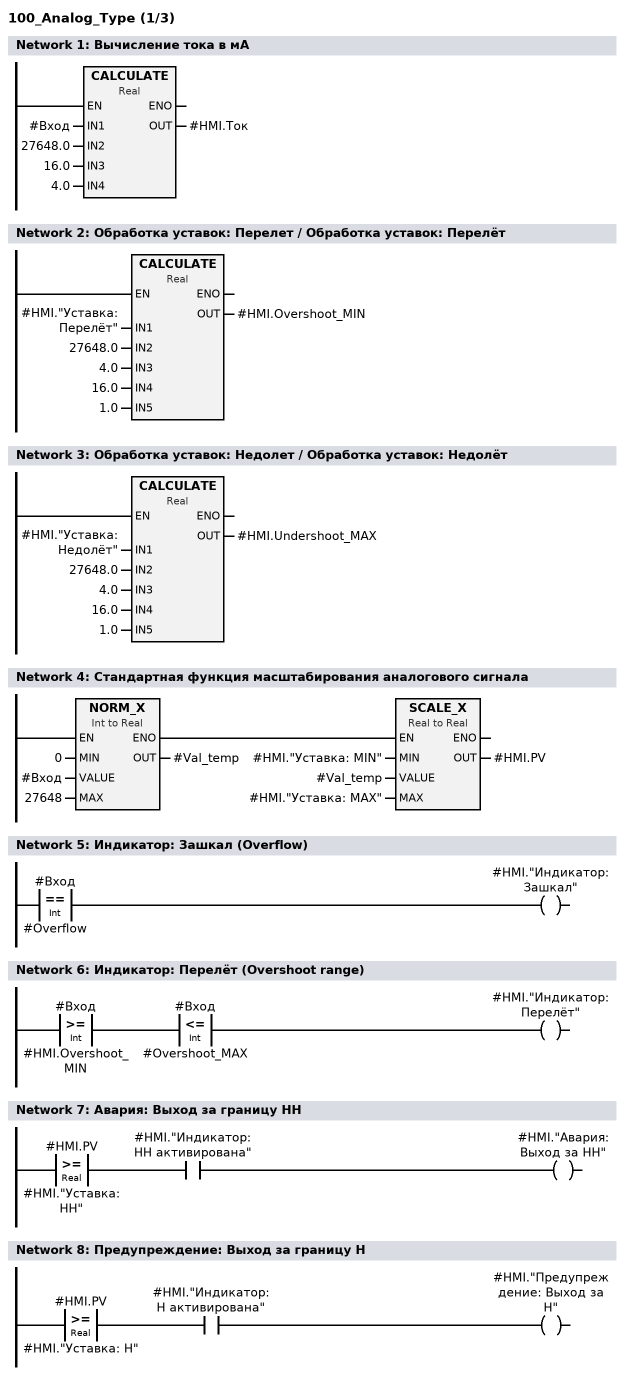
   RUNG wire#powerrail
      { S7_Templates := "SrcType := Real"; S7_Expression := "((IN3 / IN2) * IN1 + IN4)" } Calculate(in1 := #Вход, in2 := 27648.0, in3 := 16.0, in4 := 4.0, out => #HMI.Ток)
   END_RUNG
   // the same network as SCL:
   #HMI.Ток := ((16.0 / 27648.0) * #Вход + 4.0);
END_REGION

REGION Network 2: Обработка уставок: Перелет / Обработка уставок: Перелёт
   RUNG wire#powerrail
      { S7_Templates := "SrcType := Real"; S7_Expression := "((IN1- IN3) * IN2 / IN4) +IN5" } Calculate(in1 := #HMI."Уставка: Перелёт", in2 := 27648.0, in3 := 4.0, in4 := 16.0, in5 := 1.0, out => #HMI.Overshoot_MIN)
   END_RUNG
   // the same network as SCL:
   #HMI.Overshoot_MIN := ((#HMI."Уставка: Перелёт"- 4.0) * 27648.0 / 16.0) +1.0;
END_REGION

REGION Network 3: Обработка уставок: Недолет / Обработка уставок: Недолёт
   RUNG wire#powerrail
      { S7_Templates := "SrcType := Real"; S7_Expression := "((IN1- IN3) * IN2 / IN4) - IN5" } Calculate(in1 := #HMI."Уставка: Недолёт", in2 := 27648.0, in3 := 4.0, in4 := 16.0, in5 := 1.0, out => #HMI.Undershoot_MAX)
   END_RUNG
   // the same network as SCL:
   #HMI.Undershoot_MAX := ((#HMI."Уставка: Недолёт"- 4.0) * 27648.0 / 16.0) - 1.0;
END_REGION

REGION Network 4: Стандартная функция масштабирования аналогового сигнала
   RUNG wire#powerrail
      { S7_Templates := "[SrcType := Int, DestType := Real]" } Normalize(min := 0, value := #Вход, max := 27648, out => #Val_temp)
      { S7_Templates := "[SrcType := Real, DestType := Real]" } Scale(min := #HMI."Уставка: MIN", value := #Val_temp, max := #HMI."Уставка: MAX", out => #HMI.PV)
   END_RUNG
   // the same network as SCL:
   #Val_temp := NORM_X(MIN := 0, VALUE := #Вход, MAX := 27648);
   #HMI.PV := SCALE_X(MIN := #HMI."Уставка: MIN", VALUE := #Val_temp, MAX := #HMI."Уставка: MAX");
END_REGION

REGION Network 5: Индикатор: Зашкал (Overflow)
   RUNG wire#powerrail
      { S7_Templates := "SrcType := Int" } EQ_Contact(in1 := #Вход, in2 := #Overflow)
      Coil( #HMI."Индикатор: Зашкал" )
   END_RUNG
   // the same network as SCL:
   #HMI."Индикатор: Зашкал" := #Вход = #Overflow;
END_REGION

REGION Network 6: Индикатор: Перелёт (Overshoot range)
   RUNG wire#powerrail
      { S7_Templates := "SrcType := Int" } GE_Contact(in1 := #Вход, in2 := #HMI.Overshoot_MIN)
      { S7_Templates := "SrcType := Int" } LE_Contact(in1 := #Вход, in2 := #Overshoot_MAX)
      Coil( #HMI."Индикатор: Перелёт" )
   END_RUNG
   // the same network as SCL:
   #HMI."Индикатор: Перелёт" := (#Вход >= #HMI.Overshoot_MIN) AND (#Вход <= #Overshoot_MAX);
END_REGION

REGION Network 7: Авария: Выход за границу НН
   RUNG wire#powerrail
      { S7_Templates := "SrcType := Real" } GE_Contact(in1 := #HMI.PV, in2 := #HMI."Уставка: HH")
      Contact( #HMI."Индикатор: HH активирована" )
      Coil( #HMI."Авария: Выход за HH" )
   END_RUNG
   // the same network as SCL:
   #HMI."Авария: Выход за HH" := (#HMI.PV >= #HMI."Уставка: HH") AND #HMI."Индикатор: HH активирована";
END_REGION

REGION Network 8: Предупреждение: Выход за границу Н
   RUNG wire#powerrail
      { S7_Templates := "SrcType := Real" } GE_Contact(in1 := #HMI.PV, in2 := #HMI."Уставка: H")
      Contact( #HMI."Индикатор: H активирована" )
      Coil( #HMI."Предупреждение: Выход за H" )
   END_RUNG
   // the same network as SCL:
   #HMI."Предупреждение: Выход за H" := (#HMI.PV >= #HMI."Уставка: H") AND #HMI."Индикатор: H активирована";
END_REGION

REGION Network 9: Предупреждение: Выход за границу L
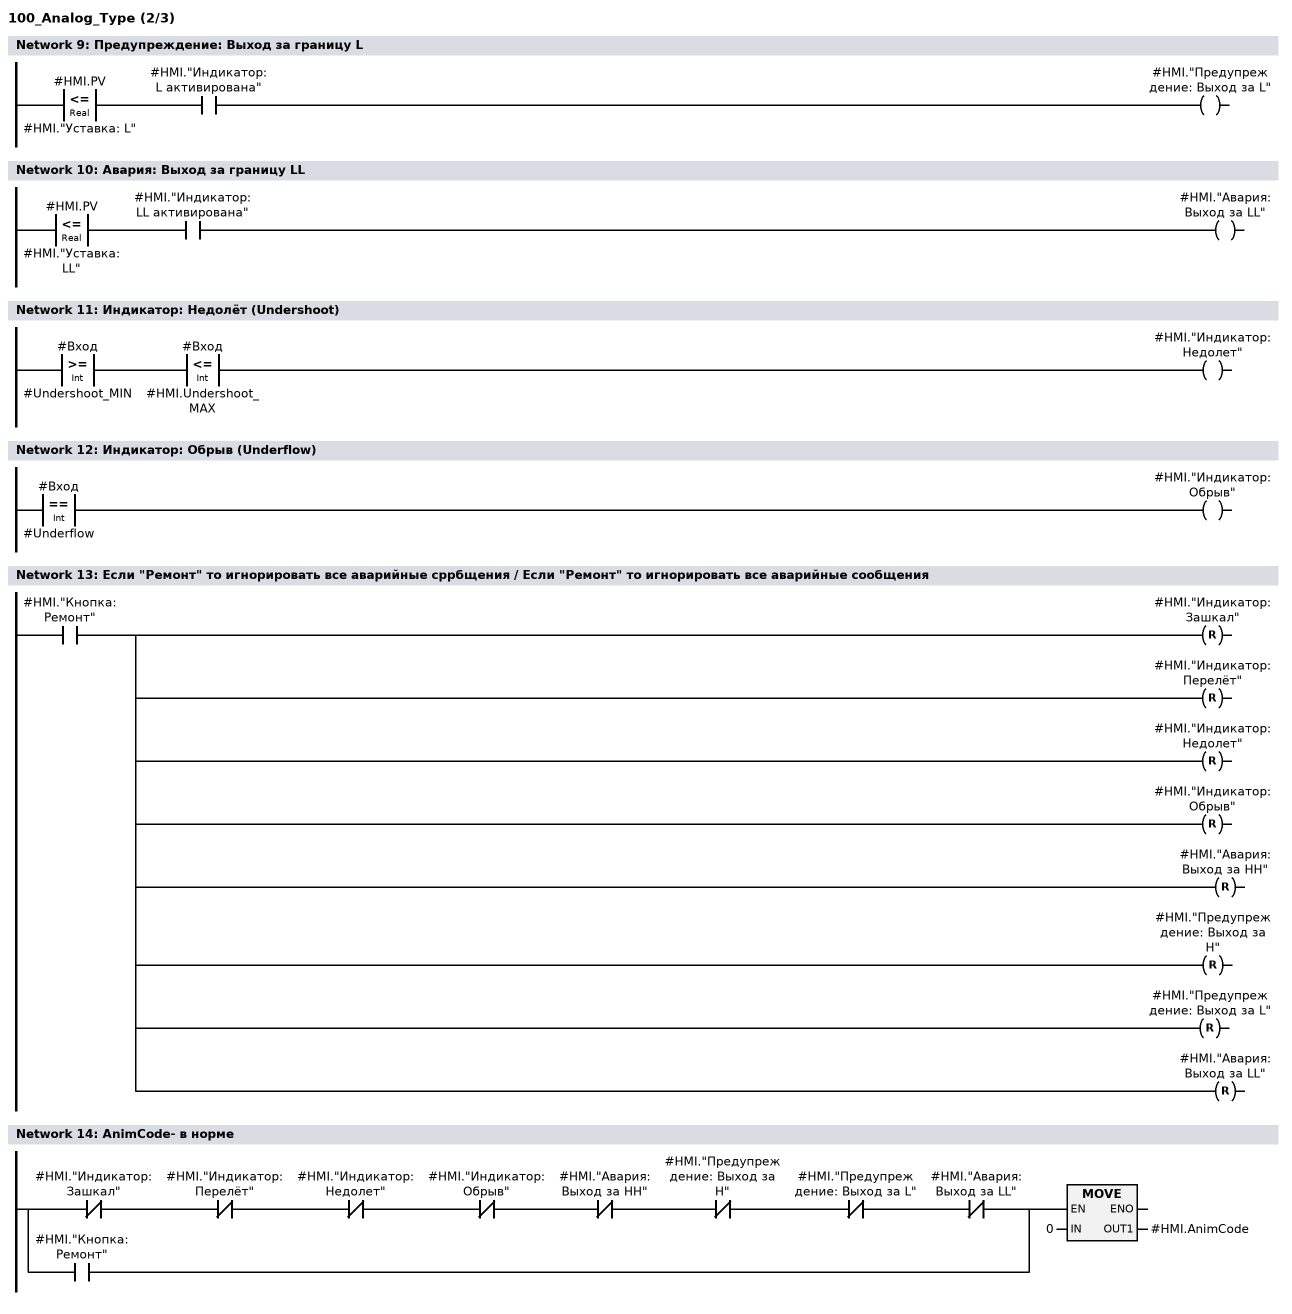
   RUNG wire#powerrail
      { S7_Templates := "SrcType := Real" } LE_Contact(in1 := #HMI.PV, in2 := #HMI."Уставка: L")
      Contact( #HMI."Индикатор: L активирована" )
      Coil( #HMI."Предупреждение: Выход за L" )
   END_RUNG
   // the same network as SCL:
   #HMI."Предупреждение: Выход за L" := (#HMI.PV <= #HMI."Уставка: L") AND #HMI."Индикатор: L активирована";
END_REGION

REGION Network 10: Авария: Выход за границу LL
   RUNG wire#powerrail
      { S7_Templates := "SrcType := Real" } LE_Contact(in1 := #HMI.PV, in2 := #HMI."Уставка: LL")
      Contact( #HMI."Индикатор: LL активирована" )
      Coil( #HMI."Авария: Выход за LL" )
   END_RUNG
   // the same network as SCL:
   #HMI."Авария: Выход за LL" := (#HMI.PV <= #HMI."Уставка: LL") AND #HMI."Индикатор: LL активирована";
END_REGION

REGION Network 11: Индикатор: Недолёт (Undershoot)
   RUNG wire#powerrail
      { S7_Templates := "SrcType := Int" } GE_Contact(in1 := #Вход, in2 := #Undershoot_MIN)
      { S7_Templates := "SrcType := Int" } LE_Contact(in1 := #Вход, in2 := #HMI.Undershoot_MAX)
      Coil( #HMI."Индикатор: Недолет" )
   END_RUNG
   // the same network as SCL:
   #HMI."Индикатор: Недолет" := (#Вход >= #Undershoot_MIN) AND (#Вход <= #HMI.Undershoot_MAX);
END_REGION

REGION Network 12: Индикатор: Обрыв (Underflow)
   RUNG wire#powerrail
      { S7_Templates := "SrcType := Int" } EQ_Contact(in1 := #Вход, in2 := #Underflow)
      Coil( #HMI."Индикатор: Обрыв" )
   END_RUNG
   // the same network as SCL:
   #HMI."Индикатор: Обрыв" := #Вход = #Underflow;
END_REGION

REGION Network 13: Если "Ремонт" то игнорировать все аварийные сррбщения / Если "Ремонт" то игнорировать все аварийные сообщения
   RUNG wire#powerrail
      Contact( #HMI."Кнопка: Ремонт" )
      wire#w1
      R_Coil( #HMI."Индикатор: Зашкал" )
   END_RUNG
   RUNG wire#w1
      R_Coil( #HMI."Индикатор: Перелёт" )
   END_RUNG
   RUNG wire#w1
      R_Coil( #HMI."Индикатор: Недолет" )
   END_RUNG
   RUNG wire#w1
      R_Coil( #HMI."Индикатор: Обрыв" )
   END_RUNG
   RUNG wire#w1
      R_Coil( #HMI."Авария: Выход за HH" )
   END_RUNG
   RUNG wire#w1
      R_Coil( #HMI."Предупреждение: Выход за H" )
   END_RUNG
   RUNG wire#w1
      R_Coil( #HMI."Предупреждение: Выход за L" )
   END_RUNG
   RUNG wire#w1
      R_Coil( #HMI."Авария: Выход за LL" )
   END_RUNG
   // the same network as SCL:
   IF #HMI."Кнопка: Ремонт" THEN
       #HMI."Индикатор: Зашкал" := FALSE;
       #HMI."Индикатор: Перелёт" := FALSE;
       #HMI."Индикатор: Недолет" := FALSE;
       #HMI."Индикатор: Обрыв" := FALSE;
       #HMI."Авария: Выход за HH" := FALSE;
       #HMI."Предупреждение: Выход за H" := FALSE;
       #HMI."Предупреждение: Выход за L" := FALSE;
       #HMI."Авария: Выход за LL" := FALSE;
   END_IF;
END_REGION

REGION Network 14: AnimCode- в норме
   RUNG wire#powerrail
      I_Contact( #HMI."Индикатор: Зашкал" )
      I_Contact( #HMI."Индикатор: Перелёт" )
      I_Contact( #HMI."Индикатор: Недолет" )
      I_Contact( #HMI."Индикатор: Обрыв" )
      I_Contact( #HMI."Авария: Выход за HH" )
      I_Contact( #HMI."Предупреждение: Выход за H" )
      I_Contact( #HMI."Предупреждение: Выход за L" )
      I_Contact( #HMI."Авария: Выход за LL" )
      wire#w1
      Move(in := 0, out1 => #HMI.AnimCode)
   END_RUNG
   RUNG wire#powerrail
      Contact( #HMI."Кнопка: Ремонт" )
   END_RUNG wire#w1
   // the same network as SCL:
   IF (NOT #HMI."Индикатор: Зашкал" AND NOT #HMI."Индикатор: Перелёт" AND NOT #HMI."Индикатор: Недолет" AND NOT #HMI."Индикатор: Обрыв" AND NOT #HMI."Авария: Выход за HH" AND NOT #HMI."Предупреждение: Выход за H" AND NOT #HMI."Предупреждение: Выход за L" AND NOT #HMI."Авария: Выход за LL") OR #HMI."Кнопка: Ремонт" THEN
       #HMI.AnimCode := 0;
   END_IF;
END_REGION

REGION Network 15: AnimCode- предупреждение
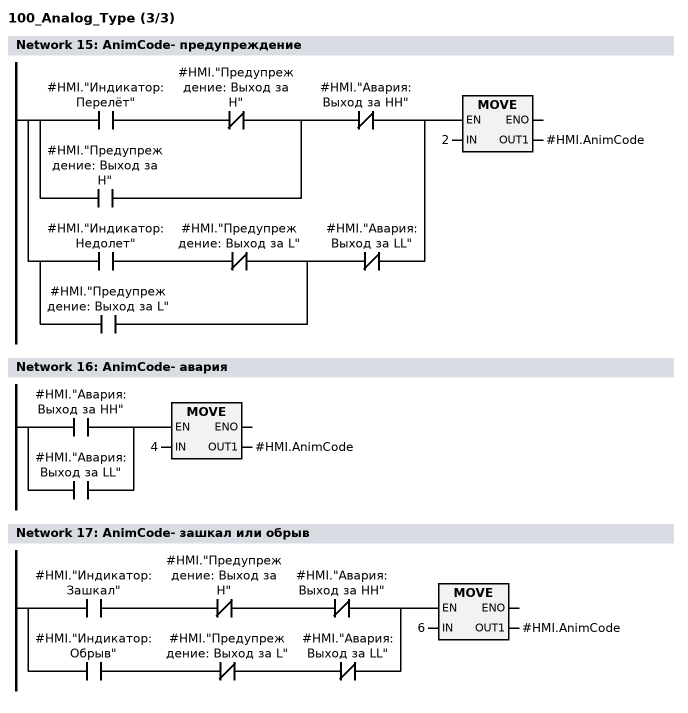
   RUNG wire#powerrail
      Contact( #HMI."Индикатор: Перелёт" )
      I_Contact( #HMI."Предупреждение: Выход за H" )
      wire#w1
      I_Contact( #HMI."Авария: Выход за HH" )
      wire#w2
      Move(in := 2, out1 => #HMI.AnimCode)
   END_RUNG
   RUNG wire#powerrail
      Contact( #HMI."Предупреждение: Выход за H" )
   END_RUNG wire#w1
   RUNG wire#powerrail
      Contact( #HMI."Индикатор: Недолет" )
      I_Contact( #HMI."Предупреждение: Выход за L" )
      wire#w3
      I_Contact( #HMI."Авария: Выход за LL" )
   END_RUNG wire#w2
   RUNG wire#powerrail
      Contact( #HMI."Предупреждение: Выход за L" )
   END_RUNG wire#w3
   // the same network as SCL:
   IF (((#HMI."Индикатор: Перелёт" AND NOT #HMI."Предупреждение: Выход за H") OR #HMI."Предупреждение: Выход за H") AND NOT #HMI."Авария: Выход за HH") OR (((#HMI."Индикатор: Недолет" AND NOT #HMI."Предупреждение: Выход за L") OR #HMI."Предупреждение: Выход за L") AND NOT #HMI."Авария: Выход за LL") THEN
       #HMI.AnimCode := 2;
   END_IF;
END_REGION

REGION Network 16: AnimCode- авария
   RUNG wire#powerrail
      Contact( #HMI."Авария: Выход за HH" )
      wire#w1
      Move(in := 4, out1 => #HMI.AnimCode)
   END_RUNG
   RUNG wire#powerrail
      Contact( #HMI."Авария: Выход за LL" )
   END_RUNG wire#w1
   // the same network as SCL:
   IF #HMI."Авария: Выход за HH" OR #HMI."Авария: Выход за LL" THEN #HMI.AnimCode := 4; END_IF;
END_REGION

REGION Network 17: AnimCode- зашкал или обрыв
   RUNG wire#powerrail
      Contact( #HMI."Индикатор: Зашкал" )
      I_Contact( #HMI."Предупреждение: Выход за H" )
      I_Contact( #HMI."Авария: Выход за HH" )
      wire#w1
      Move(in := 6, out1 => #HMI.AnimCode)
   END_RUNG
   RUNG wire#powerrail
      Contact( #HMI."Индикатор: Обрыв" )
      I_Contact( #HMI."Предупреждение: Выход за L" )
      I_Contact( #HMI."Авария: Выход за LL" )
   END_RUNG wire#w1
   // the same network as SCL:
   IF (#HMI."Индикатор: Зашкал" AND NOT #HMI."Предупреждение: Выход за H" AND NOT #HMI."Авария: Выход за HH") OR (#HMI."Индикатор: Обрыв" AND NOT #HMI."Предупреждение: Выход за L" AND NOT #HMI."Авария: Выход за LL") THEN
       #HMI.AnimCode := 6;
   END_IF;
END_REGION
END_FUNCTION

FUNCTION "101_Motor_Type" : Void   // FC101, LAD
{ S7_Optimized_Access := 'TRUE' }
VERSION : 0.1
   VAR_INPUT
      Start : Bool;
      PlcMode : Bool;
      LocalMode : Bool;
      Contactor : Bool;
      StartPulse : Bool;
      Sec_pulse : Bool;
   END_VAR
   VAR_OUTPUT
      Output : Bool;
   END_VAR
   VAR_IN_OUT
      TimeOutAccMotor : Int;
      TimeOutPreMotor : Int;
      TimeOutAccKey : Int;
      TimeOutPreKey : Int;
      ResetAlr : Bool;
      AnimCodeMotor : Int;
      AnimCodeKey : Int;
      WorkTime : DInt;
      ResetWorkTime : Bool;
   END_VAR
   VAR_TEMP
      bitTemp : Bool;
      StartTemp : Bool;
      outputt : Bool;
   END_VAR
   VAR_TEMP   // added for the SCL form of the ladder/FBD networks
      _w1 : Bool;
      _w2 : Bool;
      _w3 : Bool;
      _w4 : Bool;
      _w5 : Bool;
      _w6 : Bool;
      _w7 : Bool;
      _w8 : Bool;
   END_VAR
BEGIN

REGION Network 1
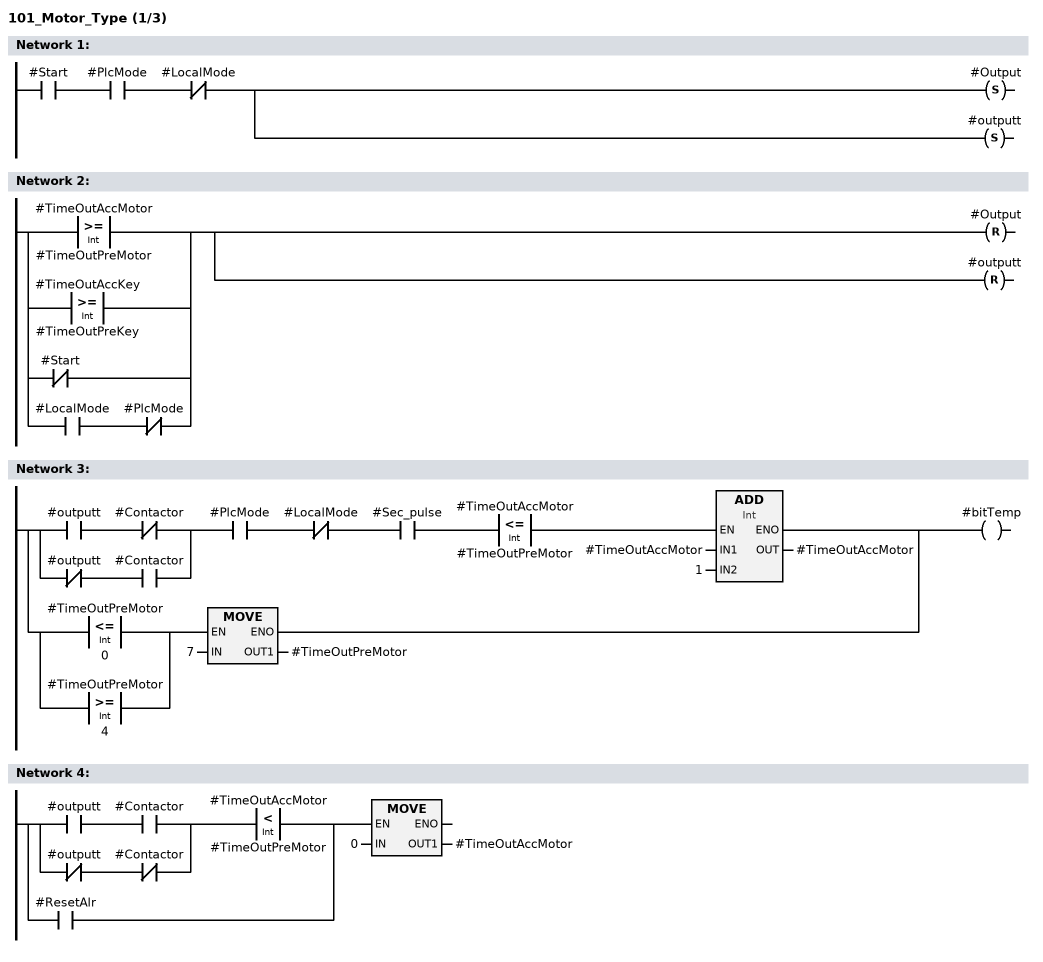
   RUNG wire#powerrail
      Contact( #Start )
      Contact( #PlcMode )
      I_Contact( #LocalMode )
      wire#w1
      S_Coil( #Output )
   END_RUNG
   RUNG wire#w1
      S_Coil( #outputt )
   END_RUNG
   // the same network as SCL:
   IF #Start AND #PlcMode AND NOT #LocalMode THEN
       #Output := TRUE;
       #outputt := TRUE;
   END_IF;
END_REGION

REGION Network 2
   RUNG wire#powerrail
      { S7_Templates := "SrcType := Int" } GE_Contact(in1 := #TimeOutAccMotor, in2 := #TimeOutPreMotor)
      wire#w1
      R_Coil( #Output )
   END_RUNG
   RUNG wire#powerrail
      { S7_Templates := "SrcType := Int" } GE_Contact(in1 := #TimeOutAccKey, in2 := #TimeOutPreKey)
   END_RUNG wire#w1
   RUNG wire#powerrail
      I_Contact( #Start )
   END_RUNG wire#w1
   RUNG wire#powerrail
      Contact( #LocalMode )
      I_Contact( #PlcMode )
   END_RUNG wire#w1
   RUNG wire#w1
      R_Coil( #outputt )
   END_RUNG
   // the same network as SCL:
   IF (#TimeOutAccMotor >= #TimeOutPreMotor) OR (#TimeOutAccKey >= #TimeOutPreKey) OR NOT #Start OR (#LocalMode AND NOT #PlcMode) THEN
       #Output := FALSE;
       #outputt := FALSE;
   END_IF;
END_REGION

REGION Network 3
   RUNG wire#powerrail
      Contact( #outputt )
      I_Contact( #Contactor )
      wire#w1
      Contact( #PlcMode )
      I_Contact( #LocalMode )
      Contact( #Sec_pulse )
      { S7_Templates := "SrcType := Int" } LE_Contact(in1 := #TimeOutAccMotor, in2 := #TimeOutPreMotor)
      { S7_Templates := "SrcType := Int"; S7_GenerateENO := "TRUE" } Add(in1 := #TimeOutAccMotor, in2 := 1, out => #TimeOutAccMotor)
      wire#w2
      Coil( #bitTemp )
   END_RUNG
   RUNG wire#powerrail
      I_Contact( #outputt )
      Contact( #Contactor )
   END_RUNG wire#w1
   RUNG wire#powerrail
      { S7_Templates := "SrcType := Int" } LE_Contact(in1 := #TimeOutPreMotor, in2 := 0)
      wire#w3
      { S7_GenerateENO := "TRUE" } Move(in := 7, out1 => #TimeOutPreMotor)
   END_RUNG wire#w2
   RUNG wire#powerrail
      { S7_Templates := "SrcType := Int" } GE_Contact(in1 := #TimeOutPreMotor, in2 := 4)
   END_RUNG wire#w3
   // the same network as SCL:
   // ENO of a box is taken as its EN; it also drops when the box reports an error
   #_w1 := ((#outputt AND NOT #Contactor) OR (NOT #outputt AND #Contactor)) AND #PlcMode AND NOT #LocalMode AND #Sec_pulse AND (#TimeOutAccMotor <= #TimeOutPreMotor);
   IF #_w1 THEN #TimeOutAccMotor := #TimeOutAccMotor + 1; END_IF;
   #_w2 := (#TimeOutPreMotor <= 0) OR (#TimeOutPreMotor >= 4);
   IF #_w2 THEN #TimeOutPreMotor := 7; END_IF;
   #bitTemp := #_w1 OR #_w2;
END_REGION

REGION Network 4
   RUNG wire#powerrail
      Contact( #outputt )
      Contact( #Contactor )
      wire#w1
      { S7_Templates := "SrcType := Int" } LT_Contact(in1 := #TimeOutAccMotor, in2 := #TimeOutPreMotor)
      wire#w2
      { S7_GenerateENO := "TRUE" } Move(in := 0, out1 => #TimeOutAccMotor)
   END_RUNG
   RUNG wire#powerrail
      I_Contact( #outputt )
      I_Contact( #Contactor )
   END_RUNG wire#w1
   RUNG wire#powerrail
      Contact( #ResetAlr )
   END_RUNG wire#w2
   // the same network as SCL:
   IF (((#outputt AND #Contactor) OR (NOT #outputt AND NOT #Contactor)) AND (#TimeOutAccMotor < #TimeOutPreMotor)) OR #ResetAlr THEN
       #TimeOutAccMotor := 0;
   END_IF;
END_REGION

REGION Network 5
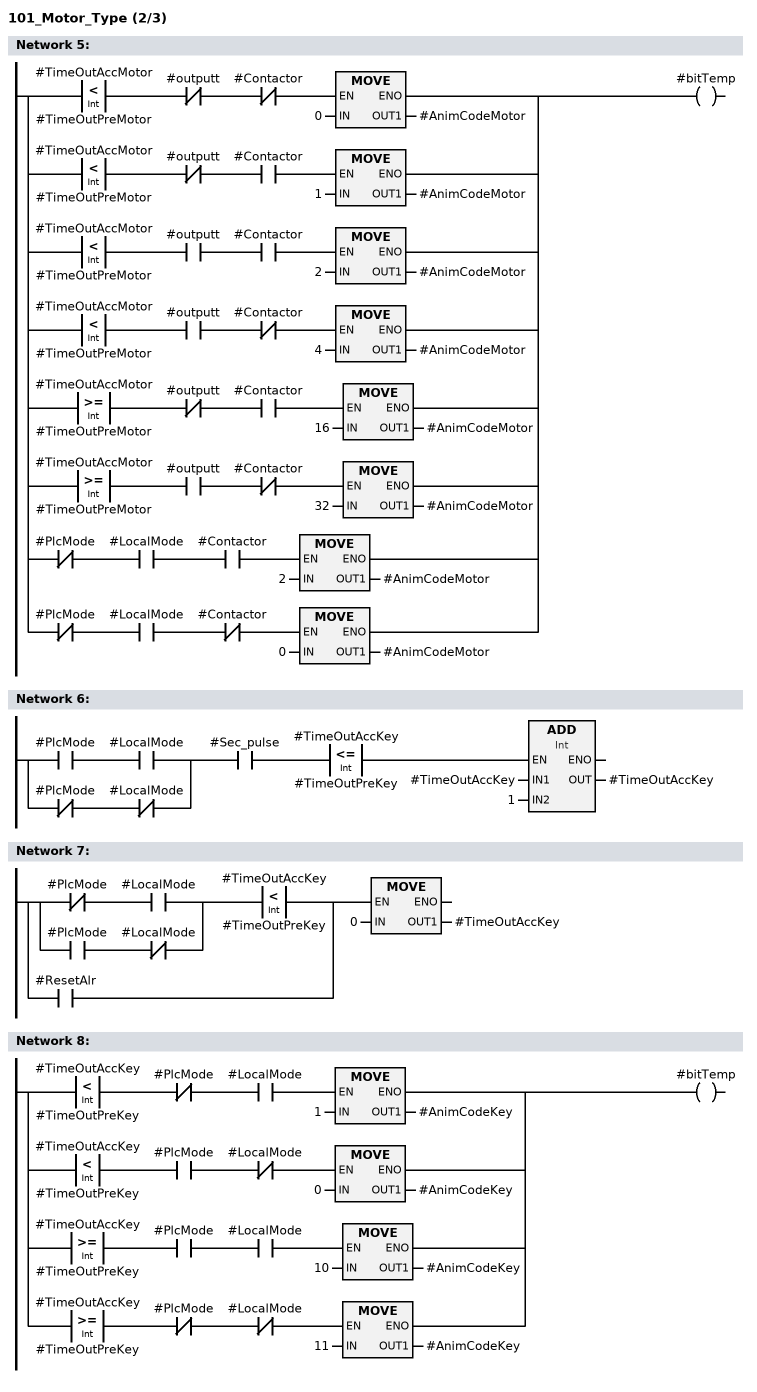
   RUNG wire#powerrail
      { S7_Templates := "SrcType := Int" } LT_Contact(in1 := #TimeOutAccMotor, in2 := #TimeOutPreMotor)
      I_Contact( #outputt )
      I_Contact( #Contactor )
      { S7_GenerateENO := "TRUE" } Move(in := 0, out1 => #AnimCodeMotor)
      wire#w1
      Coil( #bitTemp )
   END_RUNG
   RUNG wire#powerrail
      { S7_Templates := "SrcType := Int" } LT_Contact(in1 := #TimeOutAccMotor, in2 := #TimeOutPreMotor)
      I_Contact( #outputt )
      Contact( #Contactor )
      { S7_GenerateENO := "TRUE" } Move(in := 1, out1 => #AnimCodeMotor)
   END_RUNG wire#w1
   RUNG wire#powerrail
      { S7_Templates := "SrcType := Int" } LT_Contact(in1 := #TimeOutAccMotor, in2 := #TimeOutPreMotor)
      Contact( #outputt )
      Contact( #Contactor )
      { S7_GenerateENO := "TRUE" } Move(in := 2, out1 => #AnimCodeMotor)
   END_RUNG wire#w1
   RUNG wire#powerrail
      { S7_Templates := "SrcType := Int" } LT_Contact(in1 := #TimeOutAccMotor, in2 := #TimeOutPreMotor)
      Contact( #outputt )
      I_Contact( #Contactor )
      { S7_GenerateENO := "TRUE" } Move(in := 4, out1 => #AnimCodeMotor)
   END_RUNG wire#w1
   RUNG wire#powerrail
      { S7_Templates := "SrcType := Int" } GE_Contact(in1 := #TimeOutAccMotor, in2 := #TimeOutPreMotor)
      I_Contact( #outputt )
      Contact( #Contactor )
      { S7_GenerateENO := "TRUE" } Move(in := 16, out1 => #AnimCodeMotor)
   END_RUNG wire#w1
   RUNG wire#powerrail
      { S7_Templates := "SrcType := Int" } GE_Contact(in1 := #TimeOutAccMotor, in2 := #TimeOutPreMotor)
      Contact( #outputt )
      I_Contact( #Contactor )
      { S7_GenerateENO := "TRUE" } Move(in := 32, out1 => #AnimCodeMotor)
   END_RUNG wire#w1
   RUNG wire#powerrail
      I_Contact( #PlcMode )
      Contact( #LocalMode )
      Contact( #Contactor )
      { S7_GenerateENO := "TRUE" } Move(in := 2, out1 => #AnimCodeMotor)
   END_RUNG wire#w1
   RUNG wire#powerrail
      I_Contact( #PlcMode )
      Contact( #LocalMode )
      I_Contact( #Contactor )
      { S7_GenerateENO := "TRUE" } Move(in := 0, out1 => #AnimCodeMotor)
   END_RUNG wire#w1
   // the same network as SCL:
   // ENO of a box is taken as its EN; it also drops when the box reports an error
   #_w1 := (#TimeOutAccMotor < #TimeOutPreMotor) AND NOT #outputt AND NOT #Contactor;
   IF #_w1 THEN #AnimCodeMotor := 0; END_IF;
   #_w2 := (#TimeOutAccMotor < #TimeOutPreMotor) AND NOT #outputt AND #Contactor;
   IF #_w2 THEN #AnimCodeMotor := 1; END_IF;
   #_w3 := (#TimeOutAccMotor < #TimeOutPreMotor) AND #outputt AND #Contactor;
   IF #_w3 THEN #AnimCodeMotor := 2; END_IF;
   #_w4 := (#TimeOutAccMotor < #TimeOutPreMotor) AND #outputt AND NOT #Contactor;
   IF #_w4 THEN #AnimCodeMotor := 4; END_IF;
   #_w5 := (#TimeOutAccMotor >= #TimeOutPreMotor) AND NOT #outputt AND #Contactor;
   IF #_w5 THEN #AnimCodeMotor := 16; END_IF;
   #_w6 := (#TimeOutAccMotor >= #TimeOutPreMotor) AND #outputt AND NOT #Contactor;
   IF #_w6 THEN #AnimCodeMotor := 32; END_IF;
   #_w7 := NOT #PlcMode AND #LocalMode AND #Contactor;
   IF #_w7 THEN #AnimCodeMotor := 2; END_IF;
   #_w8 := NOT #PlcMode AND #LocalMode AND NOT #Contactor;
   IF #_w8 THEN #AnimCodeMotor := 0; END_IF;
   #bitTemp := #_w1 OR #_w2 OR #_w3 OR #_w4 OR #_w5 OR #_w6 OR #_w7 OR #_w8;
END_REGION

REGION Network 6
   RUNG wire#powerrail
      Contact( #PlcMode )
      Contact( #LocalMode )
      wire#w1
      Contact( #Sec_pulse )
      { S7_Templates := "SrcType := Int" } LE_Contact(in1 := #TimeOutAccKey, in2 := #TimeOutPreKey)
      { S7_Templates := "SrcType := Int"; S7_GenerateENO := "TRUE" } Add(in1 := #TimeOutAccKey, in2 := 1, out => #TimeOutAccKey)
   END_RUNG
   RUNG wire#powerrail
      I_Contact( #PlcMode )
      I_Contact( #LocalMode )
   END_RUNG wire#w1
   // the same network as SCL:
   IF ((#PlcMode AND #LocalMode) OR (NOT #PlcMode AND NOT #LocalMode)) AND #Sec_pulse AND (#TimeOutAccKey <= #TimeOutPreKey) THEN
       #TimeOutAccKey := #TimeOutAccKey + 1;
   END_IF;
END_REGION

REGION Network 7
   RUNG wire#powerrail
      I_Contact( #PlcMode )
      Contact( #LocalMode )
      wire#w1
      { S7_Templates := "SrcType := Int" } LT_Contact(in1 := #TimeOutAccKey, in2 := #TimeOutPreKey)
      wire#w2
      { S7_GenerateENO := "TRUE" } Move(in := 0, out1 => #TimeOutAccKey)
   END_RUNG
   RUNG wire#powerrail
      Contact( #PlcMode )
      I_Contact( #LocalMode )
   END_RUNG wire#w1
   RUNG wire#powerrail
      Contact( #ResetAlr )
   END_RUNG wire#w2
   // the same network as SCL:
   IF (((NOT #PlcMode AND #LocalMode) OR (#PlcMode AND NOT #LocalMode)) AND (#TimeOutAccKey < #TimeOutPreKey)) OR #ResetAlr THEN
       #TimeOutAccKey := 0;
   END_IF;
END_REGION

REGION Network 8
   RUNG wire#powerrail
      { S7_Templates := "SrcType := Int" } LT_Contact(in1 := #TimeOutAccKey, in2 := #TimeOutPreKey)
      I_Contact( #PlcMode )
      Contact( #LocalMode )
      { S7_GenerateENO := "TRUE" } Move(in := 1, out1 => #AnimCodeKey)
      wire#w1
      Coil( #bitTemp )
   END_RUNG
   RUNG wire#powerrail
      { S7_Templates := "SrcType := Int" } LT_Contact(in1 := #TimeOutAccKey, in2 := #TimeOutPreKey)
      Contact( #PlcMode )
      I_Contact( #LocalMode )
      { S7_GenerateENO := "TRUE" } Move(in := 0, out1 => #AnimCodeKey)
   END_RUNG wire#w1
   RUNG wire#powerrail
      { S7_Templates := "SrcType := Int" } GE_Contact(in1 := #TimeOutAccKey, in2 := #TimeOutPreKey)
      Contact( #PlcMode )
      Contact( #LocalMode )
      { S7_GenerateENO := "TRUE" } Move(in := 10, out1 => #AnimCodeKey)
   END_RUNG wire#w1
   RUNG wire#powerrail
      { S7_Templates := "SrcType := Int" } GE_Contact(in1 := #TimeOutAccKey, in2 := #TimeOutPreKey)
      I_Contact( #PlcMode )
      I_Contact( #LocalMode )
      { S7_GenerateENO := "TRUE" } Move(in := 11, out1 => #AnimCodeKey)
   END_RUNG wire#w1
   // the same network as SCL:
   // ENO of a box is taken as its EN; it also drops when the box reports an error
   #_w1 := (#TimeOutAccKey < #TimeOutPreKey) AND NOT #PlcMode AND #LocalMode;
   IF #_w1 THEN #AnimCodeKey := 1; END_IF;
   #_w2 := (#TimeOutAccKey < #TimeOutPreKey) AND #PlcMode AND NOT #LocalMode;
   IF #_w2 THEN #AnimCodeKey := 0; END_IF;
   #_w3 := (#TimeOutAccKey >= #TimeOutPreKey) AND #PlcMode AND #LocalMode;
   IF #_w3 THEN #AnimCodeKey := 10; END_IF;
   #_w4 := (#TimeOutAccKey >= #TimeOutPreKey) AND NOT #PlcMode AND NOT #LocalMode;
   IF #_w4 THEN #AnimCodeKey := 11; END_IF;
   #bitTemp := #_w1 OR #_w2 OR #_w3 OR #_w4;
END_REGION

REGION Network 9
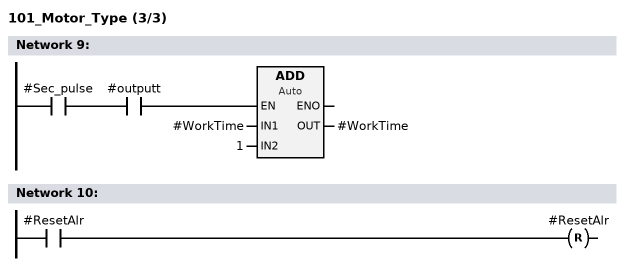
   RUNG wire#powerrail
      Contact( #Sec_pulse )
      Contact( #outputt )
      Add(in1 := #WorkTime, in2 := 1, out => #WorkTime)
   END_RUNG
   // the same network as SCL:
   IF #Sec_pulse AND #outputt THEN #WorkTime := #WorkTime + 1; END_IF;
END_REGION

REGION Network 10
   RUNG wire#powerrail
      Contact( #ResetAlr )
      R_Coil( #ResetAlr )
   END_RUNG
   // the same network as SCL:
   IF #ResetAlr THEN #ResetAlr := FALSE; END_IF;
END_REGION
END_FUNCTION

FUNCTION "102_Discret_Type" : Void   // FC102, LAD
{ S7_Optimized_Access := 'FALSE' }
VERSION : 0.1
   VAR_INPUT
      INPUT : Bool;
   END_VAR
   VAR_OUTPUT
      OUT_BOOL : Bool;
      OUT_INT : Int;
   END_VAR
BEGIN

REGION Network 1
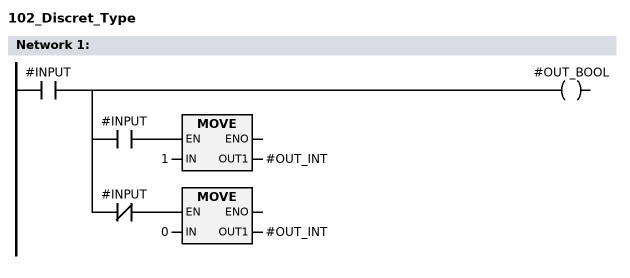
   RUNG wire#powerrail
      Contact( #INPUT )
      wire#w1
      Coil( #OUT_BOOL )
   END_RUNG
   RUNG wire#w1
      Contact( #INPUT )
      { S7_GenerateENO := "TRUE" } Move(in := 1, out1 => #OUT_INT)
   END_RUNG
   RUNG wire#w1
      I_Contact( #INPUT )
      { S7_GenerateENO := "TRUE" } Move(in := 0, out1 => #OUT_INT)
   END_RUNG
   // the same network as SCL:
   #OUT_BOOL := #INPUT;
   IF #INPUT AND #INPUT THEN #OUT_INT := 1; END_IF;
   IF #INPUT AND NOT #INPUT THEN #OUT_INT := 0; END_IF;
END_REGION
END_FUNCTION

FUNCTION "104_FC_Narabotka" : Void   // FC104, SCL
{ S7_Optimized_Access := 'TRUE' }
VERSION : 0.1
   VAR_INPUT
      Puls_Second : Bool;
   END_VAR
   VAR_IN_OUT
      t : "Narabotki";
   END_VAR
BEGIN
       IF #Puls_Second AND #t.old = 0 THEN
           #t.Second := #t.Second + 1;
           IF #t.Second >= 60 THEN
               #t.Second := 0;
               #t.Minute := #t.Minute + 1;
               IF #t.Minute >= 60 THEN
                   #t.Minute := 0;
                   #t.Hour := #t.Hour + 1;
               END_IF;
           END_IF;
           #t.old := 1;
       END_IF;

   IF #Puls_Second = 0 AND #t.old THEN
       #t.old := 0;
   END_IF;

   IF #t.reset THEN
       #t.Hour := 0;
       #t.Minute := 0;
       #t.Second := 0;
   END_IF;
END_FUNCTION

FUNCTION "105_Valve_Type" : Void   // FC105, FBD
{ S7_Optimized_Access := 'FALSE' }
VERSION : 0.1
   VAR_INPUT
      PLC_Mode : Bool;
      Local_Mode : Bool;
      SwOpen : Bool;
      SwClose : Bool;
      CmdOpen : Bool;
      CmdClose : Bool;
      Sec_pulse : Bool;
   END_VAR
   VAR_OUTPUT
      OutputOpen : Bool;   // Открытие
      OutputClose : Bool;   // Закрытие
   END_VAR
   VAR_IN_OUT
      ResetALr : Bool;   // Сброс нарушения
      ResetWorkTime : Bool;   // Сброс часов работы мотора
      TimeOutPreValve : Int;
      TimeOutAccValve : Int;
      TimeOutPreKey : Int;
      TimeOutAccKey : Int;
      WorkTime : DInt;
      AnimCodeValve : Int;   // Код анимации крана
      AnimCodeKey : Int;   // Код анимации ключа Сблокированный/Ручной
      OpenPulse : Bool;
      ClosePulse : Bool;
   END_VAR
   VAR_TEMP
      Starttemp : Bool;
      bitTemp : Bool;
      OpenWithoutCmd : Bool;
      CloseWithoutCmd : Bool;
      TempOpenPulse : Bool;
      TempClosePulse : Bool;
   END_VAR
   VAR_TEMP   // added for the SCL form of the ladder/FBD networks
      _w1 : Bool;
      _w2 : Bool;
      _w3 : Bool;
      _w4 : Bool;
   END_VAR
BEGIN

REGION Network 1: Открытие крана